
REGION Network 14: Ni100 RTD sensor type
   RUNG wire#powerrail
      { S7_Templates := "SrcType := Int" } EQ_Contact(in1 := #iInSensorType, in2 := "IoScaling.S7Analog.Types.Ni100")
      wire#w1
      { S7_GenerateENO := "TRUE" } Move(in := "IoScaling.S7Analog.Ni100.iRawMin", out1 => #iRawMin)
      { S7_GenerateENO := "TRUE" } Move(in := "IoScaling.S7Analog.Ni100.iRawMax", out1 => #iRawMax)
   END_RUNG
   RUNG wire#w1
      { S7_GenerateENO := "TRUE" } Move(in := "IoScaling.S7Analog.Ni100.rScaledMin", out1 => #rScaledMin)
      { S7_GenerateENO := "TRUE" } Move(in := "IoScaling.S7Analog.Ni100.rScaledMax", out1 => #rScaledMax)
   END_RUNG
   // the same network as SCL:
   // ENO of a box is taken as its EN; it also drops when the box reports an error
   IF #iInSensorType = "IoScaling.S7Analog.Types.Ni100" THEN
       #iRawMin := "IoScaling.S7Analog.Ni100.iRawMin";
       #iRawMax := "IoScaling.S7Analog.Ni100.iRawMax";
       #rScaledMin := "IoScaling.S7Analog.Ni100.rScaledMin";
       #rScaledMax := "IoScaling.S7Analog.Ni100.rScaledMax";
   END_IF;
END_REGION

REGION Network 15: Ni100 Climate RTD sensor type
   RUNG wire#powerrail
      { S7_Templates := "SrcType := Int" } EQ_Contact(in1 := #iInSensorType, in2 := "IoScaling.S7Analog.Types.Ni100.Climate")
      wire#w1
      { S7_GenerateENO := "TRUE" } Move(in := "IoScaling.S7Analog.Ni100.Climate.iRawMin", out1 => #iRawMin)
      { S7_GenerateENO := "TRUE" } Move(in := "IoScaling.S7Analog.Ni100.Climate.iRawMax", out1 => #iRawMax)
   END_RUNG
   RUNG wire#w1
      { S7_GenerateENO := "TRUE" } Move(in := "IoScaling.S7Analog.Ni100.Climate.rScaledMin", out1 => #rScaledMin)
      { S7_GenerateENO := "TRUE" } Move(in := "IoScaling.S7Analog.Ni100.Climate.rScaledMax", out1 => #rScaledMax)
   END_RUNG
   // the same network as SCL:
   // ENO of a box is taken as its EN; it also drops when the box reports an error
   IF #iInSensorType = "IoScaling.S7Analog.Types.Ni100.Climate" THEN
       #iRawMin := "IoScaling.S7Analog.Ni100.Climate.iRawMin";
       #iRawMax := "IoScaling.S7Analog.Ni100.Climate.iRawMax";
       #rScaledMin := "IoScaling.S7Analog.Ni100.Climate.rScaledMin";
       #rScaledMax := "IoScaling.S7Analog.Ni100.Climate.rScaledMax";
   END_IF;
END_REGION

REGION Network 16: --------------------------------------------------------- Errors ------------------------------------------------------------------
END_REGION

REGION Network 17: Error: High high alarm
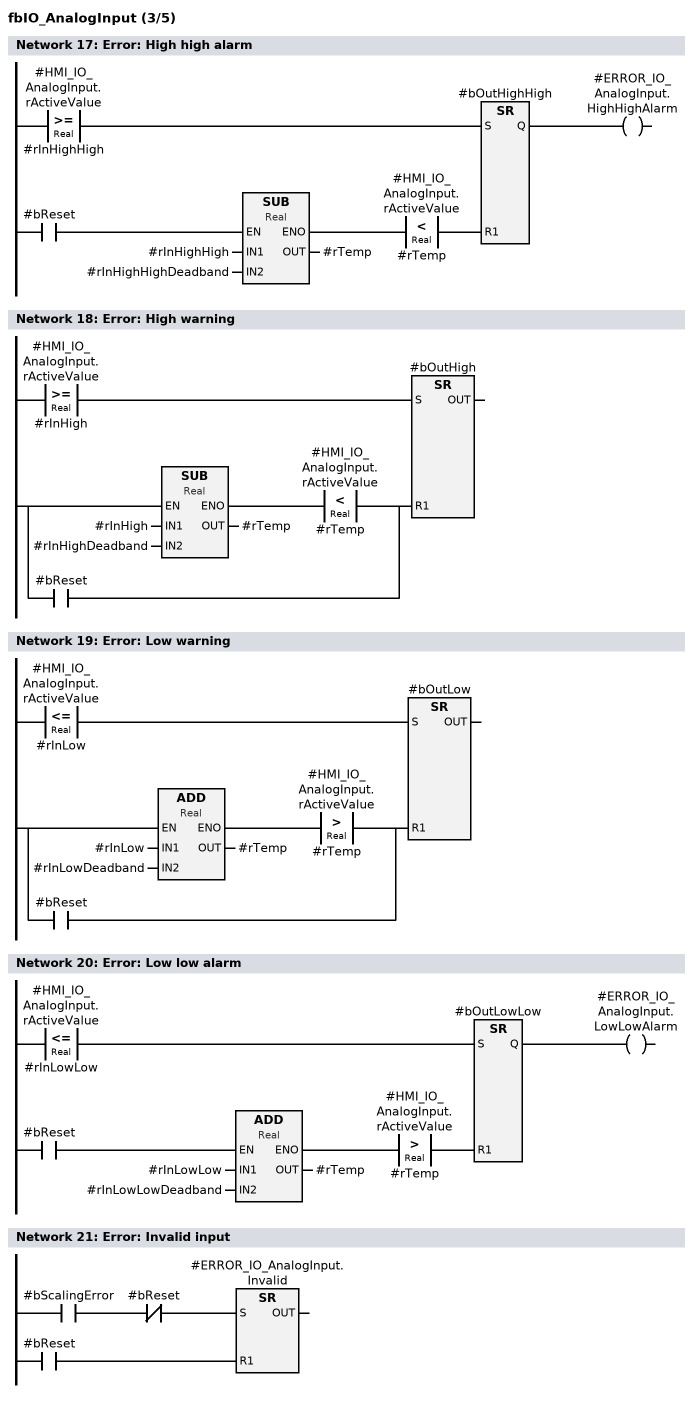
   RUNG wire#powerrail
      { S7_Templates := "SrcType := Real" } GE_Contact(in1 := #HMI_IO_AnalogInput.rActiveValue, in2 := #rInHighHigh)
      S_SR(operand := #bOutHighHigh, r1 := wire#w1)
      Coil( #ERROR_IO_AnalogInput.HighHighAlarm )
   END_RUNG
   RUNG wire#powerrail
      Contact( #bReset )
      { S7_Templates := "SrcType := Real"; S7_GenerateENO := "TRUE" } Sub(in1 := #rInHighHigh, in2 := #rInHighHighDeadband, out => #rTemp)
      { S7_Templates := "SrcType := Real" } LT_Contact(in1 := #HMI_IO_AnalogInput.rActiveValue, in2 := #rTemp)
   END_RUNG wire#w1
   // the same network as SCL:
   // ENO of a box is taken as its EN; it also drops when the box reports an error
   IF #bReset THEN #rTemp := #rInHighHigh - #rInHighHighDeadband; END_IF;
   IF #HMI_IO_AnalogInput.rActiveValue >= #rInHighHigh THEN
       #bOutHighHigh := TRUE;   // SR flip-flop
   END_IF;
   IF #bReset AND (#HMI_IO_AnalogInput.rActiveValue < #rTemp) THEN #bOutHighHigh := FALSE; END_IF;
   #ERROR_IO_AnalogInput.HighHighAlarm := #bOutHighHigh;
END_REGION

REGION Network 18: Error: High warning
   RUNG wire#powerrail
      { S7_Templates := "SrcType := Real" } GE_Contact(in1 := #HMI_IO_AnalogInput.rActiveValue, in2 := #rInHigh)
      S_SR(operand := #bOutHigh, r1 := wire#w1)
   END_RUNG
   RUNG wire#powerrail
      { S7_Templates := "SrcType := Real"; S7_GenerateENO := "TRUE" } Sub(in1 := #rInHigh, in2 := #rInHighDeadband, out => #rTemp)
      { S7_Templates := "SrcType := Real" } LT_Contact(in1 := #HMI_IO_AnalogInput.rActiveValue, in2 := #rTemp)
   END_RUNG wire#w1
   RUNG wire#powerrail
      Contact( #bReset )
   END_RUNG wire#w1
   // the same network as SCL:
   // ENO of a box is taken as its EN; it also drops when the box reports an error
   #rTemp := #rInHigh - #rInHighDeadband;
   IF #HMI_IO_AnalogInput.rActiveValue >= #rInHigh THEN
       #bOutHigh := TRUE;   // SR flip-flop
   END_IF;
   IF (#HMI_IO_AnalogInput.rActiveValue < #rTemp) OR #bReset THEN #bOutHigh := FALSE; END_IF;
END_REGION

REGION Network 19: Error: Low warning
   RUNG wire#powerrail
      { S7_Templates := "SrcType := Real" } LE_Contact(in1 := #HMI_IO_AnalogInput.rActiveValue, in2 := #rInLow)
      S_SR(operand := #bOutLow, r1 := wire#w1)
   END_RUNG
   RUNG wire#powerrail
      { S7_Templates := "SrcType := Real"; S7_GenerateENO := "TRUE" } Add(in1 := #rInLow, in2 := #rInLowDeadband, out => #rTemp)
      { S7_Templates := "SrcType := Real" } GT_Contact(in1 := #HMI_IO_AnalogInput.rActiveValue, in2 := #rTemp)
   END_RUNG wire#w1
   RUNG wire#powerrail
      Contact( #bReset )
   END_RUNG wire#w1
   // the same network as SCL:
   // ENO of a box is taken as its EN; it also drops when the box reports an error
   #rTemp := #rInLow + #rInLowDeadband;
   IF #HMI_IO_AnalogInput.rActiveValue <= #rInLow THEN
       #bOutLow := TRUE;   // SR flip-flop
   END_IF;
   IF (#HMI_IO_AnalogInput.rActiveValue > #rTemp) OR #bReset THEN #bOutLow := FALSE; END_IF;
END_REGION

REGION Network 20: Error: Low low alarm
   RUNG wire#powerrail
      { S7_Templates := "SrcType := Real" } LE_Contact(in1 := #HMI_IO_AnalogInput.rActiveValue, in2 := #rInLowLow)
      S_SR(operand := #bOutLowLow, r1 := wire#w1)
      Coil( #ERROR_IO_AnalogInput.LowLowAlarm )
   END_RUNG
   RUNG wire#powerrail
      Contact( #bReset )
      { S7_Templates := "SrcType := Real"; S7_GenerateENO := "TRUE" } Add(in1 := #rInLowLow, in2 := #rInLowLowDeadband, out => #rTemp)
      { S7_Templates := "SrcType := Real" } GT_Contact(in1 := #HMI_IO_AnalogInput.rActiveValue, in2 := #rTemp)
   END_RUNG wire#w1
   // the same network as SCL:
   // ENO of a box is taken as its EN; it also drops when the box reports an error
   IF #bReset THEN #rTemp := #rInLowLow + #rInLowLowDeadband; END_IF;
   IF #HMI_IO_AnalogInput.rActiveValue <= #rInLowLow THEN
       #bOutLowLow := TRUE;   // SR flip-flop
   END_IF;
   IF #bReset AND (#HMI_IO_AnalogInput.rActiveValue > #rTemp) THEN #bOutLowLow := FALSE; END_IF;
   #ERROR_IO_AnalogInput.LowLowAlarm := #bOutLowLow;
END_REGION

REGION Network 21: Error: Invalid input
   RUNG wire#powerrail
      Contact( #bScalingError )
      I_Contact( #bReset )
      S_SR(operand := #ERROR_IO_AnalogInput.Invalid, r1 := wire#w1)
   END_RUNG
   RUNG wire#powerrail
      Contact( #bReset )
   END_RUNG wire#w1
   // the same network as SCL:
   IF #bScalingError AND NOT #bReset THEN
       #ERROR_IO_AnalogInput.Invalid := TRUE;   // SR flip-flop
   END_IF;
   IF #bReset THEN #ERROR_IO_AnalogInput.Invalid := FALSE; END_IF;
END_REGION

REGION Network 22: Scroll errors on the HMI
   // Call the Error-Scroller which cyles through all possible errors and checks 
   // their state for display on the HMI
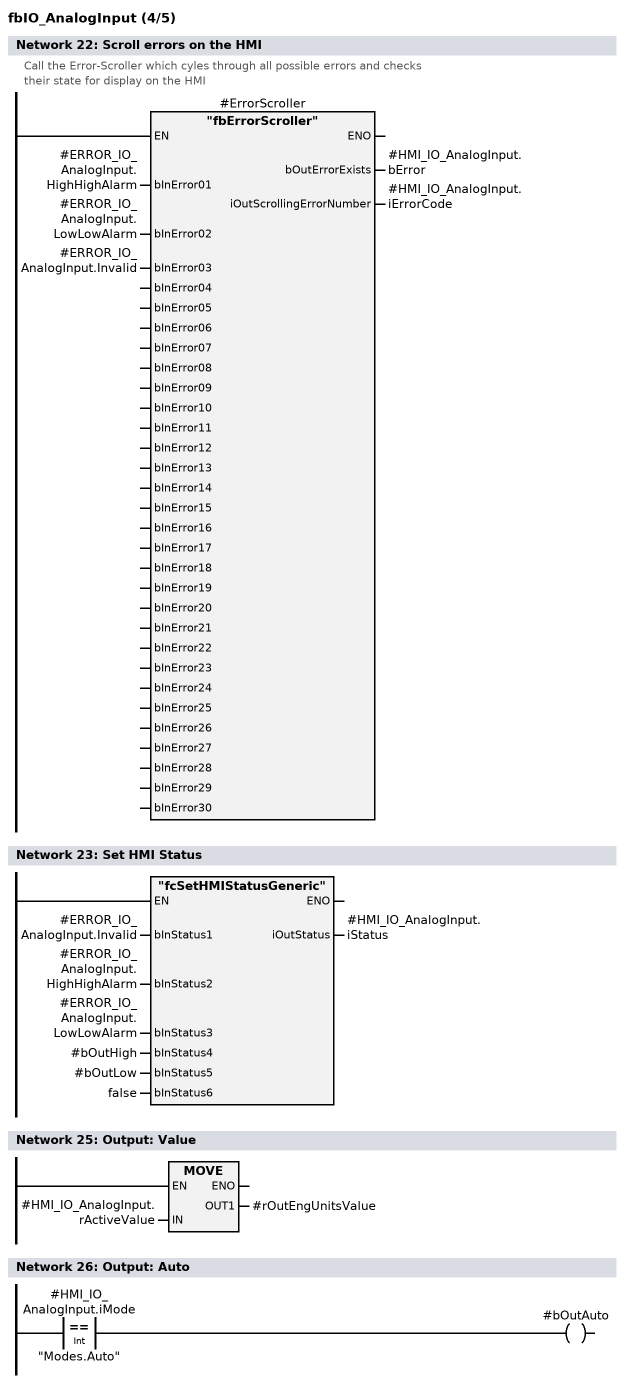
   RUNG wire#powerrail
      #ErrorScroller(bInError01 := #ERROR_IO_AnalogInput.HighHighAlarm, bInError02 := #ERROR_IO_AnalogInput.LowLowAlarm, bInError03 := #ERROR_IO_AnalogInput.Invalid, bInError04 :=, bInError05 :=, bInError06 :=, bInError07 :=, bInError08 :=, bInError09 :=, bInError10 :=, bInError11 :=, bInError12 :=, bInError13 :=, bInError14 :=, bInError15 :=, bInError16 :=, bInError17 :=, bInError18 :=, bInError19 :=, bInError20 :=, bInError21 :=, bInError22 :=, bInError23 :=, bInError24 :=, bInError25 :=, bInError26 :=, bInError27 :=, bInError28 :=, bInError29 :=, bInError30 :=, bOutErrorExists => #HMI_IO_AnalogInput.bError, iOutScrollingErrorNumber => #HMI_IO_AnalogInput.iErrorCode)
   END_RUNG
   // the same network as SCL:
   #ErrorScroller(bInError01 := #ERROR_IO_AnalogInput.HighHighAlarm,   // "fbErrorScroller"
                  bInError02 := #ERROR_IO_AnalogInput.LowLowAlarm,
                  bInError03 := #ERROR_IO_AnalogInput.Invalid,
                  bOutErrorExists => #HMI_IO_AnalogInput.bError,
                  iOutScrollingErrorNumber => #HMI_IO_AnalogInput.iErrorCode);
END_REGION

REGION Network 23: Set HMI Status
   RUNG wire#powerrail
      "fcSetHMIStatusGeneric"(bInStatus1 := #ERROR_IO_AnalogInput.Invalid, bInStatus2 := #ERROR_IO_AnalogInput.HighHighAlarm, bInStatus3 := #ERROR_IO_AnalogInput.LowLowAlarm, bInStatus4 := #bOutHigh, bInStatus5 := #bOutLow, bInStatus6 := false, iOutStatus => #HMI_IO_AnalogInput.iStatus)
   END_RUNG
   // the same network as SCL:
   "fcSetHMIStatusGeneric"(bInStatus1 := #ERROR_IO_AnalogInput.Invalid,
                           bInStatus2 := #ERROR_IO_AnalogInput.HighHighAlarm,
                           bInStatus3 := #ERROR_IO_AnalogInput.LowLowAlarm,
                           bInStatus4 := #bOutHigh,
                           bInStatus5 := #bOutLow,
                           bInStatus6 := false,
                           iOutStatus => #HMI_IO_AnalogInput.iStatus);
END_REGION

REGION Network 24: --------------------------------------------------------- Outputs ------------------------------------------------------------------
END_REGION

REGION Network 25: Output: Value
   RUNG wire#powerrail
      { S7_GenerateENO := "TRUE" } Move(in := #HMI_IO_AnalogInput.rActiveValue, out1 => #rOutEngUnitsValue)
   END_RUNG
   // the same network as SCL:
   #rOutEngUnitsValue := #HMI_IO_AnalogInput.rActiveValue;
END_REGION

REGION Network 26: Output: Auto
   RUNG wire#powerrail
      { S7_Templates := "SrcType := Int" } EQ_Contact(in1 := #HMI_IO_AnalogInput.iMode, in2 := "Modes.Auto")
      Coil( #bOutAuto )
   END_RUNG
   // the same network as SCL:
   #bOutAuto := #HMI_IO_AnalogInput.iMode = "Modes.Auto";
END_REGION

REGION Network 27: Output: Error
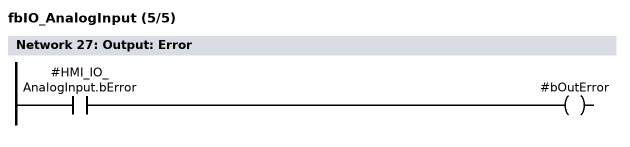
   RUNG wire#powerrail
      Contact( #HMI_IO_AnalogInput.bError )
      Coil( #bOutError )
   END_RUNG
   // the same network as SCL:
   #bOutError := #HMI_IO_AnalogInput.bError;
END_REGION
END_FUNCTION_BLOCK

FUNCTION_BLOCK "fbIO_AnalogOutput"   // FB141, LAD
TITLE = Controls an analog output
{ S7_Optimized_Access := 'FALSE' }
VERSION : 0.1
   VAR_TEMP   // added for the SCL form of the ladder/FBD networks
      _w1 : Bool;
   END_VAR
BEGIN

REGION Network 1: --------------------------------------------------------- Inputs ------------------------------------------------------------------
END_REGION

REGION Network 2: Read HMI input buttons
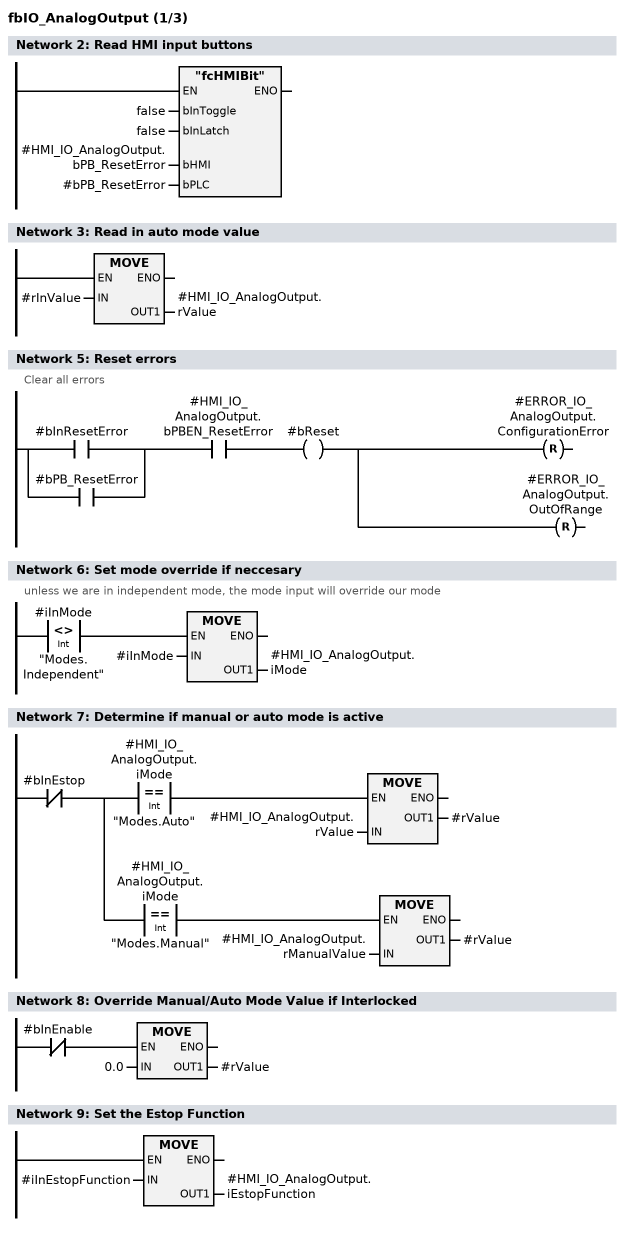
   RUNG wire#powerrail
      "fcHMIBit"(bInToggle := false, bInLatch := false, bHMI := #HMI_IO_AnalogOutput.bPB_ResetError, bPLC := #bPB_ResetError)
   END_RUNG
   // the same network as SCL:
   "fcHMIBit"(bInToggle := false,
              bInLatch := false,
              bHMI := #HMI_IO_AnalogOutput.bPB_ResetError,
              bPLC := #bPB_ResetError);
END_REGION

REGION Network 3: Read in auto mode value
   RUNG wire#powerrail
      { S7_GenerateENO := "TRUE" } Move(in := #rInValue, out1 => #HMI_IO_AnalogOutput.rValue)
   END_RUNG
   // the same network as SCL:
   #HMI_IO_AnalogOutput.rValue := #rInValue;
END_REGION

REGION Network 4: --------------------------------------------------- Control Logic ------------------------------------------------------------
END_REGION

REGION Network 5: Reset errors
   // Clear all errors
   RUNG wire#powerrail
      Contact( #bInResetError )
      wire#w1
      Contact( #HMI_IO_AnalogOutput.bPBEN_ResetError )
      Coil( #bReset )
      wire#w2
      R_Coil( #ERROR_IO_AnalogOutput.ConfigurationError )
   END_RUNG
   RUNG wire#powerrail
      Contact( #bPB_ResetError )
   END_RUNG wire#w1
   RUNG wire#w2
      R_Coil( #ERROR_IO_AnalogOutput.OutOfRange )
   END_RUNG
   // the same network as SCL:
   #bReset := (#bInResetError OR #bPB_ResetError) AND #HMI_IO_AnalogOutput.bPBEN_ResetError;
   IF #bReset THEN
       #ERROR_IO_AnalogOutput.ConfigurationError := FALSE;
       #ERROR_IO_AnalogOutput.OutOfRange := FALSE;
   END_IF;
END_REGION

REGION Network 6: Set mode override if neccesary
   // unless we are in independent mode, the mode input will override our mode
   RUNG wire#powerrail
      { S7_Templates := "SrcType := Int" } NE_Contact(in1 := #iInMode, in2 := "Modes.Independent")
      { S7_GenerateENO := "TRUE" } Move(in := #iInMode, out1 => #HMI_IO_AnalogOutput.iMode)
   END_RUNG
   // the same network as SCL:
   IF #iInMode <> "Modes.Independent" THEN #HMI_IO_AnalogOutput.iMode := #iInMode; END_IF;
END_REGION

REGION Network 7: Determine if manual or auto mode is active
   RUNG wire#powerrail
      I_Contact( #bInEstop )
      wire#w1
      { S7_Templates := "SrcType := Int" } EQ_Contact(in1 := #HMI_IO_AnalogOutput.iMode, in2 := "Modes.Auto")
      { S7_GenerateENO := "TRUE" } Move(in := #HMI_IO_AnalogOutput.rValue, out1 => #rValue)
   END_RUNG
   RUNG wire#w1
      { S7_Templates := "SrcType := Int" } EQ_Contact(in1 := #HMI_IO_AnalogOutput.iMode, in2 := "Modes.Manual")
      { S7_GenerateENO := "TRUE" } Move(in := #HMI_IO_AnalogOutput.rManualValue, out1 => #rValue)
   END_RUNG
   // the same network as SCL:
   IF NOT #bInEstop AND (#HMI_IO_AnalogOutput.iMode = "Modes.Auto") THEN
       #rValue := #HMI_IO_AnalogOutput.rValue;
   END_IF;
   IF NOT #bInEstop AND (#HMI_IO_AnalogOutput.iMode = "Modes.Manual") THEN
       #rValue := #HMI_IO_AnalogOutput.rManualValue;
   END_IF;
END_REGION

REGION Network 8: Override Manual/Auto Mode Value if Interlocked
   RUNG wire#powerrail
      I_Contact( #bInEnable )
      { S7_GenerateENO := "TRUE" } Move(in := 0.0, out1 => #rValue)
   END_RUNG
   // the same network as SCL:
   IF NOT #bInEnable THEN #rValue := 0.0; END_IF;
END_REGION

REGION Network 9: Set the Estop Function
   RUNG wire#powerrail
      Move(in := #iInEstopFunction, out1 => #HMI_IO_AnalogOutput.iEstopFunction)
   END_RUNG
   // the same network as SCL:
   #HMI_IO_AnalogOutput.iEstopFunction := #iInEstopFunction;
END_REGION

REGION Network 10: Determine E-Stop set point
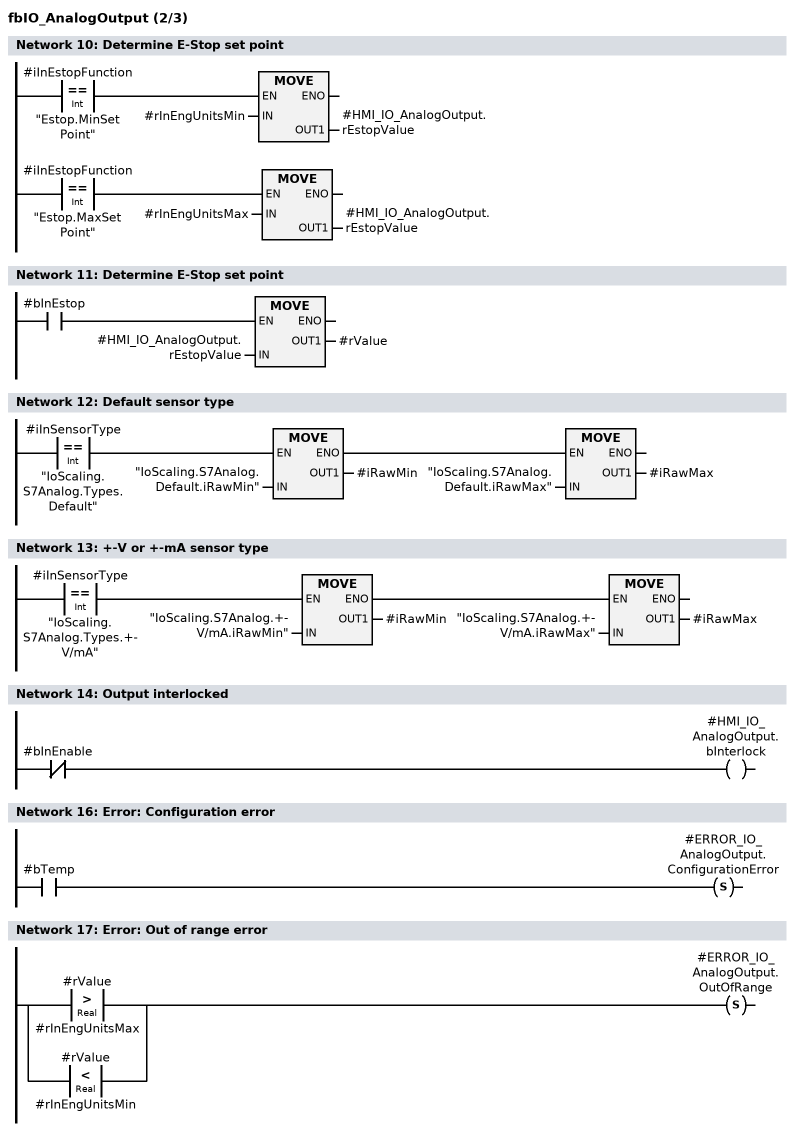
   RUNG wire#powerrail
      { S7_Templates := "SrcType := Int" } EQ_Contact(in1 := #iInEstopFunction, in2 := "Estop.MinSetPoint")
      { S7_GenerateENO := "TRUE" } Move(in := #rInEngUnitsMin, out1 => #HMI_IO_AnalogOutput.rEstopValue)
   END_RUNG
   RUNG wire#powerrail
      { S7_Templates := "SrcType := Int" } EQ_Contact(in1 := #iInEstopFunction, in2 := "Estop.MaxSetPoint")
      { S7_GenerateENO := "TRUE" } Move(in := #rInEngUnitsMax, out1 => #HMI_IO_AnalogOutput.rEstopValue)
   END_RUNG
   // the same network as SCL:
   IF #iInEstopFunction = "Estop.MinSetPoint" THEN
       #HMI_IO_AnalogOutput.rEstopValue := #rInEngUnitsMin;
   END_IF;
   IF #iInEstopFunction = "Estop.MaxSetPoint" THEN
       #HMI_IO_AnalogOutput.rEstopValue := #rInEngUnitsMax;
   END_IF;
END_REGION

REGION Network 11: Determine E-Stop set point
   RUNG wire#powerrail
      Contact( #bInEstop )
      { S7_GenerateENO := "TRUE" } Move(in := #HMI_IO_AnalogOutput.rEstopValue, out1 => #rValue)
   END_RUNG
   // the same network as SCL:
   IF #bInEstop THEN #rValue := #HMI_IO_AnalogOutput.rEstopValue; END_IF;
END_REGION

REGION Network 12: Default sensor type
   RUNG wire#powerrail
      { S7_Templates := "SrcType := Int" } EQ_Contact(in1 := #iInSensorType, in2 := "IoScaling.S7Analog.Types.Default")
      { S7_GenerateENO := "TRUE" } Move(in := "IoScaling.S7Analog.Default.iRawMin", out1 => #iRawMin)
      { S7_GenerateENO := "TRUE" } Move(in := "IoScaling.S7Analog.Default.iRawMax", out1 => #iRawMax)
   END_RUNG
   // the same network as SCL:
   // ENO of a box is taken as its EN; it also drops when the box reports an error
   IF #iInSensorType = "IoScaling.S7Analog.Types.Default" THEN
       #iRawMin := "IoScaling.S7Analog.Default.iRawMin";
       #iRawMax := "IoScaling.S7Analog.Default.iRawMax";
   END_IF;
END_REGION

REGION Network 13: +-V or +-mA sensor type
   RUNG wire#powerrail
      { S7_Templates := "SrcType := Int" } EQ_Contact(in1 := #iInSensorType, in2 := "IoScaling.S7Analog.Types.+-V/mA")
      { S7_GenerateENO := "TRUE" } Move(in := "IoScaling.S7Analog.+-V/mA.iRawMin", out1 => #iRawMin)
      { S7_GenerateENO := "TRUE" } Move(in := "IoScaling.S7Analog.+-V/mA.iRawMax", out1 => #iRawMax)
   END_RUNG
   // the same network as SCL:
   // ENO of a box is taken as its EN; it also drops when the box reports an error
   IF #iInSensorType = "IoScaling.S7Analog.Types.+-V/mA" THEN
       #iRawMin := "IoScaling.S7Analog.+-V/mA.iRawMin";
       #iRawMax := "IoScaling.S7Analog.+-V/mA.iRawMax";
   END_IF;
END_REGION

REGION Network 14: Output interlocked
   RUNG wire#powerrail
      I_Contact( #bInEnable )
      Coil( #HMI_IO_AnalogOutput.bInterlock )
   END_RUNG
   // the same network as SCL:
   #HMI_IO_AnalogOutput.bInterlock := NOT #bInEnable;
END_REGION

REGION Network 15: --------------------------------------------------------- Errors ------------------------------------------------------------------
END_REGION

REGION Network 16: Error: Configuration error
   RUNG wire#powerrail
      Contact( #bTemp )
      S_Coil( #ERROR_IO_AnalogOutput.ConfigurationError )
   END_RUNG
   // the same network as SCL:
   IF #bTemp THEN #ERROR_IO_AnalogOutput.ConfigurationError := TRUE; END_IF;
END_REGION

REGION Network 17: Error: Out of range error
   RUNG wire#powerrail
      { S7_Templates := "SrcType := Real" } GT_Contact(in1 := #rValue, in2 := #rInEngUnitsMax)
      wire#w1
      S_Coil( #ERROR_IO_AnalogOutput.OutOfRange )
   END_RUNG
   RUNG wire#powerrail
      { S7_Templates := "SrcType := Real" } LT_Contact(in1 := #rValue, in2 := #rInEngUnitsMin)
   END_RUNG wire#w1
   // the same network as SCL:
   IF (#rValue > #rInEngUnitsMax) OR (#rValue < #rInEngUnitsMin) THEN
       #ERROR_IO_AnalogOutput.OutOfRange := TRUE;
   END_IF;
END_REGION

REGION Network 18: Scroll errors on the HMI
   // Call the Error-Scroller which cyles through all possible errors and checks 
   // their state for display on the HMI
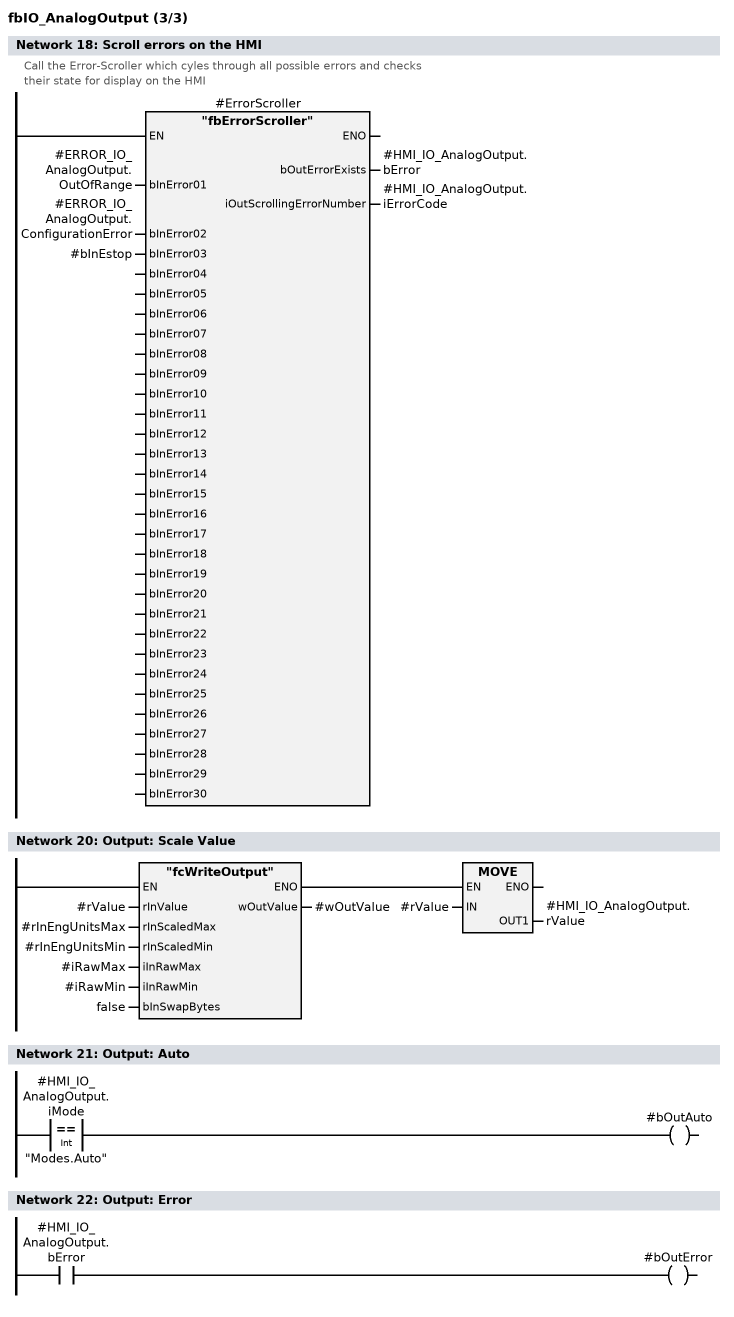
   RUNG wire#powerrail
      #ErrorScroller(bInError01 := #ERROR_IO_AnalogOutput.OutOfRange, bInError02 := #ERROR_IO_AnalogOutput.ConfigurationError, bInError03 := #bInEstop, bInError04 :=, bInError05 :=, bInError06 :=, bInError07 :=, bInError08 :=, bInError09 :=, bInError10 :=, bInError11 :=, bInError12 :=, bInError13 :=, bInError14 :=, bInError15 :=, bInError16 :=, bInError17 :=, bInError18 :=, bInError19 :=, bInError20 :=, bInError21 :=, bInError22 :=, bInError23 :=, bInError24 :=, bInError25 :=, bInError26 :=, bInError27 :=, bInError28 :=, bInError29 :=, bInError30 :=, bOutErrorExists => #HMI_IO_AnalogOutput.bError, iOutScrollingErrorNumber => #HMI_IO_AnalogOutput.iErrorCode)
   END_RUNG
   // the same network as SCL:
   #ErrorScroller(bInError01 := #ERROR_IO_AnalogOutput.OutOfRange,   // "fbErrorScroller"
                  bInError02 := #ERROR_IO_AnalogOutput.ConfigurationError,
                  bInError03 := #bInEstop,
                  bOutErrorExists => #HMI_IO_AnalogOutput.bError,
                  iOutScrollingErrorNumber => #HMI_IO_AnalogOutput.iErrorCode);
END_REGION

REGION Network 19: --------------------------------------------------------- Outputs ------------------------------------------------------------------
END_REGION

REGION Network 20: Output: Scale Value
   RUNG wire#powerrail
      "fcWriteOutput"(rInValue := #rValue, rInScaledMax := #rInEngUnitsMax, rInScaledMin := #rInEngUnitsMin, iInRawMax := #iRawMax, iInRawMin := #iRawMin, bInSwapBytes := false, wOutValue => #wOutValue)
      Move(in := #rValue, out1 => #HMI_IO_AnalogOutput.rValue)
   END_RUNG
   // the same network as SCL:
   "fcWriteOutput"(rInValue := #rValue,
                   rInScaledMax := #rInEngUnitsMax,
                   rInScaledMin := #rInEngUnitsMin,
                   iInRawMax := #iRawMax,
                   iInRawMin := #iRawMin,
                   bInSwapBytes := false,
                   wOutValue => #wOutValue,
                   ENO => #_w1);
   IF #_w1 THEN #HMI_IO_AnalogOutput.rValue := #rValue; END_IF;
END_REGION

REGION Network 21: Output: Auto
   RUNG wire#powerrail
      { S7_Templates := "SrcType := Int" } EQ_Contact(in1 := #HMI_IO_AnalogOutput.iMode, in2 := "Modes.Auto")
      Coil( #bOutAuto )
   END_RUNG
   // the same network as SCL:
   #bOutAuto := #HMI_IO_AnalogOutput.iMode = "Modes.Auto";
END_REGION

REGION Network 22: Output: Error
   RUNG wire#powerrail
      Contact( #HMI_IO_AnalogOutput.bError )
      Coil( #bOutError )
   END_RUNG
   // the same network as SCL:
   #bOutError := #HMI_IO_AnalogOutput.bError;
END_REGION
END_FUNCTION_BLOCK

// folder: Library Blocks/Process

FUNCTION_BLOCK "fbInterlock"   // FB160, LAD
TITLE = Compiles interlock conditions for a system
{ S7_Optimized_Access := 'FALSE' }
VERSION : 0.1
BEGIN

REGION Network 1: Determine interlock status
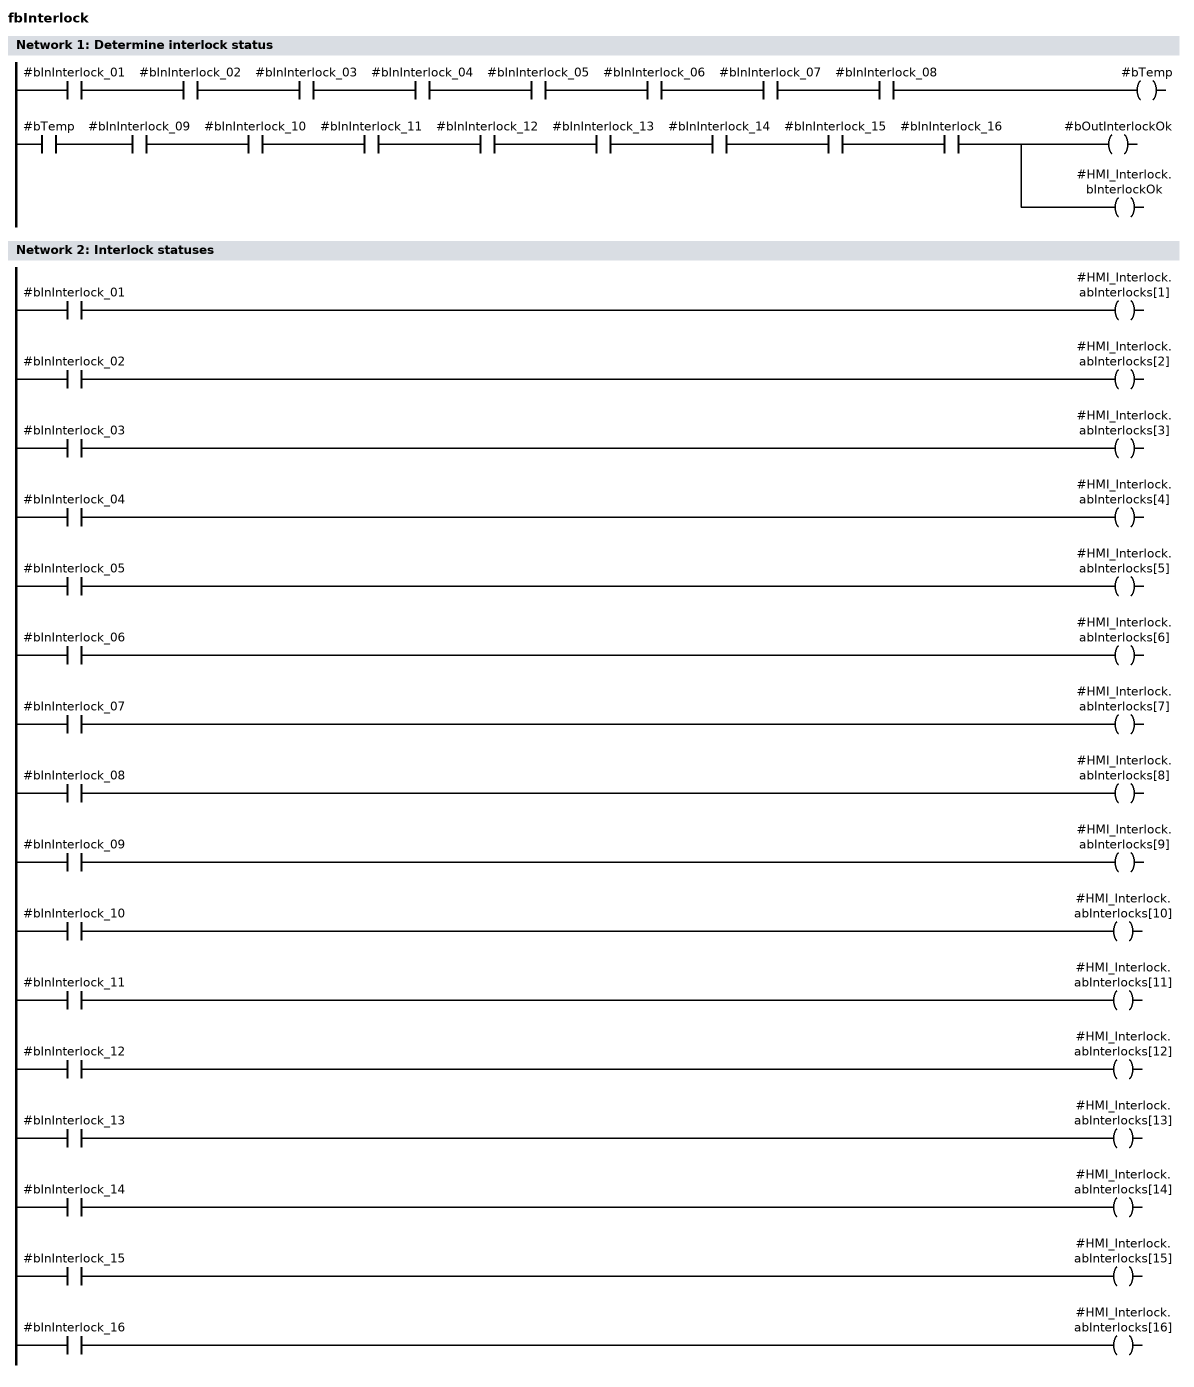
   RUNG wire#powerrail
      Contact( #bInInterlock_01 )
      Contact( #bInInterlock_02 )
      Contact( #bInInterlock_03 )
      Contact( #bInInterlock_04 )
      Contact( #bInInterlock_05 )
      Contact( #bInInterlock_06 )
      Contact( #bInInterlock_07 )
      Contact( #bInInterlock_08 )
      Coil( #bTemp )
   END_RUNG
   RUNG wire#powerrail
      Contact( #bTemp )
      Contact( #bInInterlock_09 )
      Contact( #bInInterlock_10 )
      Contact( #bInInterlock_11 )
      Contact( #bInInterlock_12 )
      Contact( #bInInterlock_13 )
      Contact( #bInInterlock_14 )
      Contact( #bInInterlock_15 )
      Contact( #bInInterlock_16 )
      wire#w1
      Coil( #bOutInterlockOk )
   END_RUNG
   RUNG wire#w1
      Coil( #HMI_Interlock.bInterlockOk )
   END_RUNG
   // the same network as SCL:
   #bTemp := #bInInterlock_01 AND #bInInterlock_02 AND #bInInterlock_03 AND #bInInterlock_04 AND #bInInterlock_05 AND #bInInterlock_06 AND #bInInterlock_07 AND #bInInterlock_08;
   #bOutInterlockOk := #bTemp AND #bInInterlock_09 AND #bInInterlock_10 AND #bInInterlock_11 AND #bInInterlock_12 AND #bInInterlock_13 AND #bInInterlock_14 AND #bInInterlock_15 AND #bInInterlock_16;
   #HMI_Interlock.bInterlockOk := #bOutInterlockOk;
END_REGION

REGION Network 2: Interlock statuses
   RUNG wire#powerrail
      Contact( #bInInterlock_01 )
      Coil( #HMI_Interlock.abInterlocks[1] )
   END_RUNG
   RUNG wire#powerrail
      Contact( #bInInterlock_02 )
      Coil( #HMI_Interlock.abInterlocks[2] )
   END_RUNG
   RUNG wire#powerrail
      Contact( #bInInterlock_03 )
      Coil( #HMI_Interlock.abInterlocks[3] )
   END_RUNG
   RUNG wire#powerrail
      Contact( #bInInterlock_04 )
      Coil( #HMI_Interlock.abInterlocks[4] )
   END_RUNG
   RUNG wire#powerrail
      Contact( #bInInterlock_05 )
      Coil( #HMI_Interlock.abInterlocks[5] )
   END_RUNG
   RUNG wire#powerrail
      Contact( #bInInterlock_06 )
      Coil( #HMI_Interlock.abInterlocks[6] )
   END_RUNG
   RUNG wire#powerrail
      Contact( #bInInterlock_07 )
      Coil( #HMI_Interlock.abInterlocks[7] )
   END_RUNG
   RUNG wire#powerrail
      Contact( #bInInterlock_08 )
      Coil( #HMI_Interlock.abInterlocks[8] )
   END_RUNG
   RUNG wire#powerrail
      Contact( #bInInterlock_09 )
      Coil( #HMI_Interlock.abInterlocks[9] )
   END_RUNG
   RUNG wire#powerrail
      Contact( #bInInterlock_10 )
      Coil( #HMI_Interlock.abInterlocks[10] )
   END_RUNG
   RUNG wire#powerrail
      Contact( #bInInterlock_11 )
      Coil( #HMI_Interlock.abInterlocks[11] )
   END_RUNG
   RUNG wire#powerrail
      Contact( #bInInterlock_12 )
      Coil( #HMI_Interlock.abInterlocks[12] )
   END_RUNG
   RUNG wire#powerrail
      Contact( #bInInterlock_13 )
      Coil( #HMI_Interlock.abInterlocks[13] )
   END_RUNG
   RUNG wire#powerrail
      Contact( #bInInterlock_14 )
      Coil( #HMI_Interlock.abInterlocks[14] )
   END_RUNG
   RUNG wire#powerrail
      Contact( #bInInterlock_15 )
      Coil( #HMI_Interlock.abInterlocks[15] )
   END_RUNG
   RUNG wire#powerrail
      Contact( #bInInterlock_16 )
      Coil( #HMI_Interlock.abInterlocks[16] )
   END_RUNG
   // the same network as SCL:
   #HMI_Interlock.abInterlocks[1] := #bInInterlock_01;
   #HMI_Interlock.abInterlocks[2] := #bInInterlock_02;
   #HMI_Interlock.abInterlocks[3] := #bInInterlock_03;
   #HMI_Interlock.abInterlocks[4] := #bInInterlock_04;
   #HMI_Interlock.abInterlocks[5] := #bInInterlock_05;
   #HMI_Interlock.abInterlocks[6] := #bInInterlock_06;
   #HMI_Interlock.abInterlocks[7] := #bInInterlock_07;
   #HMI_Interlock.abInterlocks[8] := #bInInterlock_08;
   #HMI_Interlock.abInterlocks[9] := #bInInterlock_09;
   #HMI_Interlock.abInterlocks[10] := #bInInterlock_10;
   #HMI_Interlock.abInterlocks[11] := #bInInterlock_11;
   #HMI_Interlock.abInterlocks[12] := #bInInterlock_12;
   #HMI_Interlock.abInterlocks[13] := #bInInterlock_13;
   #HMI_Interlock.abInterlocks[14] := #bInInterlock_14;
   #HMI_Interlock.abInterlocks[15] := #bInInterlock_15;
   #HMI_Interlock.abInterlocks[16] := #bInInterlock_16;
END_REGION
END_FUNCTION_BLOCK

FUNCTION_BLOCK "fbAlarmWarning"   // FB161, LAD
TITLE = Controls a latching alarm
{ S7_Optimized_Access := 'FALSE' }
VERSION : 0.1
BEGIN

REGION Network 1: Set warning condition
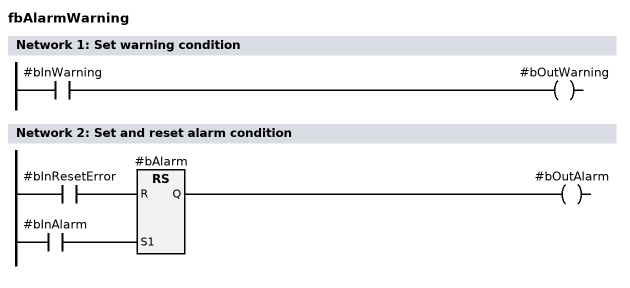
   RUNG wire#powerrail
      Contact( #bInWarning )
      Coil( #bOutWarning )
   END_RUNG
   // the same network as SCL:
   #bOutWarning := #bInWarning;
END_REGION

REGION Network 2: Set and reset alarm condition
   RUNG wire#powerrail
      Contact( #bInResetError )
      S_RS(operand := #bAlarm, s1 := wire#w1)
      Coil( #bOutAlarm )
   END_RUNG
   RUNG wire#powerrail
      Contact( #bInAlarm )
   END_RUNG wire#w1
   // the same network as SCL:
   IF #bInResetError THEN
       #bAlarm := FALSE;   // RS flip-flop
   END_IF;
   IF #bInAlarm THEN #bAlarm := TRUE; END_IF;
   #bOutAlarm := #bAlarm;
END_REGION
END_FUNCTION_BLOCK

FUNCTION_BLOCK "fbPID_CompactInterface"   // FB165, LAD
TITLE = Controls and interfacs with a PID_Compact object
{ S7_Optimized_Access := 'FALSE' }
VERSION : 0.1
   VAR_TEMP   // added for the SCL form of the ladder/FBD networks
      _w1 : Bool;
      _w2 : Bool;
      _w3 : Bool;
      _w4 : Bool;
      _w5 : Bool;
   END_VAR
BEGIN

REGION Network 1: --------------------------------------------------------- Inputs ------------------------------------------------------------------
END_REGION

REGION Network 2: Read HMI input buttons
